           IF #statBatteryFamily1 = 16#0A THEN
               #HMI.State.Details.batFamily := 1;          //BAT1600
           ELSIF #statBatteryFamily1 = 16#09 THEN
               IF #statBatteryFamily2 = 16#07 THEN
                   #HMI.State.Details.batFamily := 3;          //Third Party Battery
               ELSE
                   #HMI.State.Details.batFamily := 2;          //UPS1100
               END_IF;
           END_IF;
           #HMI.State.batteryType := #statDataBatteryInfo.batteryDetails[0].batteryType;
           #HMI.State.endOfChargeVolt := INT_TO_REAL(#statDataBatteryInfo.batteryDetails[0].eocv) * 0.01;
           FOR #tempIterator := 0 TO 5 BY 1 DO
               #HMI.State.batteryDetails[#tempIterator].batteryLEDState := #statDataBatteryInfo.batteryDetails[#tempIterator].batLEDState;
               #HMI.State.batteryDetails[#tempIterator].batteryOpState := #statDataBatteryInfo.batteryDetails[#tempIterator].batOpState;
               #HMI.State.batteryDetails[#tempIterator].batteryCalcHealth := #statDataBatteryInfo.batteryDetails[#tempIterator].batCalcHealth;
           END_FOR;
           #HMI.State.chargingOpState := #statDataStateInfo.chargingOpState;
           // Cyclic Data
           #HMI.Mode.bufferMode := #statCyclicData[1];
           #HMI.Mode.readyForBuffering := #statCyclicData[2];
           #HMI.State.batteryChargeLevel := #statCyclicData[6];
           #statCyclicCount := 1;
       END_IF;

       //if Buffer_mode = 255, start Timer
       IF #HMI.Mode.bufferMode = 255 AND NOT #statBlockTimer AND NOT #statSetTimer THEN
           #statSetTimer := 1;
       END_IF;

       IF #HMI.Mode.bufferMode = 0 THEN
           #statSetTimer := 0;
           #statCmdDone := FALSE;
           #statBlockTimer := 0;
       END_IF;

       //BlockTimer - block
       #statTimerObj(IN := #statSetTimer,   // IN: BOOL
                     PT := #statBufferTime); // IN: TIME

       //Timer "Reset signal"
       IF #statTimerObj.Q = 1 THEN
           //if time elapse > UPS_ready_for_reset = 1
           #upsReadyForReset := 1;
           #statSetTimer := 0;
           #statBlockTimer := 1;
       END_IF;

       //reset UPS_ready_for_reset = 0 / set command parameter
       IF #upsExecuteReset = 1 AND NOT #statWrReq AND (#statBlockTimer = TRUE) AND (#statCmdDone = FALSE) THEN
           #statWrReq := 1;
           #statDataUPSCmd.commandID := 8207; //Command Remote Reset
           #statDataUPSCmd.parameter1 := INT_TO_BYTE(#statDataBufParam.bufferTime2);
           #statDataUPSCmd.parameter2 := #statDataResetParam;   //Parameter
           #upsReadyForReset := 0;
       END_IF;

       //write UPS Command
       #statDataRecordWrite(REQ := #statWrReq, ID := #addrIn, INDEX := 16, LEN := 4, RECORD := #statDataUPSCmd);

       IF #statDataRecordWrite.DONE OR #statDataRecordWrite.ERROR THEN
           #statWrReq := 0;
       END_IF;

       IF #statDataRecordWrite.DONE THEN
           #statCmdDone := TRUE;
       END_IF;

       // char to string > Order_number
       Chars_TO_Strg(Chars := #statDataDeviceInfo.orderNumber, pChars := 0, Cnt := 0, Strg => #statOrderNumberStr);
       #HMI.State.Details.orderNumber := #statOrderNumberStr;

       // char to string > Serial_number
       Chars_TO_Strg(Chars := #statDataDeviceInfo.serialNumber, pChars := 0, Cnt := 0, Strg => #statSerialNumberStr);
       #HMI.State.Details.serialNumber := #statSerialNumberStr;

       // char to string > Device_name
       Chars_TO_Strg(Chars := #statDataDeviceInfo.deviceName, pChars := 0, Cnt := 0, Strg => #statDeviceNameStr);
       #HMI.State.Details.deviceName := #statDeviceNameStr;

       // char to string > Version_number
       Chars_TO_Strg(Chars := #statDataDeviceInfo.versionNumber, pChars := 0, Cnt := 0, Strg => #statVersionNumberStr);
       #HMI.State.Details.versionNumber := #statVersionNumberStr;

       IF #statRetVal <> 0 AND #statCyclicCount = 1 THEN
           //setting acyclic data to default values
           #HMI.State.Details.orderNumber := ' ';
           #HMI.State.Details.serialNumber := ' ';
           #HMI.State.Details.deviceName := ' ';
           #HMI.State.Details.versionNumber := ' ';
           #HMI.State.Details.deviceHwRevision := 0;
           #HMI.State.Details.deviceSwRevision3 := 0;
           #HMI.State.Details.deviceSwRevision2 := 0;
           #HMI.State.Details.deviceSwRevision1 := 0;
           #HMI.State.numOfBatteries := 0;
           #HMI.State.Details.batFamily := 0;
           #HMI.State.batteryType := 0;
           #upsReadyForReset := 0;
       END_IF;
   END_IF;
END_REGION
END_FUNCTION_BLOCK

// folder: 1}Library/Analog

FUNCTION_BLOCK "Average"   // FB12, LAD
{ S7_Optimized_Access := 'TRUE' }
VERSION : 0.1
   VAR_INPUT
      TX1 : Real;
      TX2 : Real;
   END_VAR
   VAR_OUTPUT
      SAI : Real;
   END_VAR
BEGIN

REGION Network 1
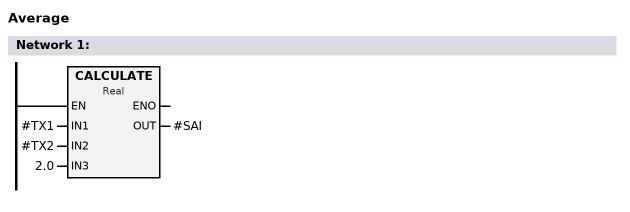
   RUNG wire#powerrail
      { S7_Templates := "SrcType := Real"; S7_Expression := "(IN1+IN2)/IN3" } Calculate(in1 := #TX1, in2 := #TX2, in3 := 2.0, out => #SAI)
   END_RUNG
   // the same network as SCL:
   #SAI := (#TX1+#TX2)/2.0;
END_REGION
END_FUNCTION_BLOCK

FUNCTION_BLOCK "AI Monitor"   // FB19, SCL
TITLE = Analog Input Monitor
{ S7_Optimized_Access := 'TRUE' }
AUTHOR : JLopez
VERSION : 0.1
// Monitor up to 6 Analog Inputs and execute AVG, in Range, deviation.
   VAR_INPUT
      "Enable Block" : Bool;   // Enable Block Execution
      "AI Num" : Int;   // Numbers of Analog Inputs Max: 6
      AvgSP : Real;   // Average SP Furnace Temperature
      "Min Range" : Real;   // Minimum Furnace Temperature Range
      "Max Range" : Real;   // Maximun Furnace Temperature Range
      MinAvgValue : Real := 0.0;   // Min Average Hysteresis Range
      MaxAvgValue : Real := 0.0;   // Max Average Hysteresis Range
      EnableDeviationMon : Bool;
      AlarmDeviation : Real := 25.0;
      MaxDeviation : Real := 50.0;   // Maximun deviation Allows
      MaxAboveTemp : Real := 50.0;
   END_VAR
   VAR_IN_OUT
      Avg : Real;   // Average Value
      AvgReached : Bool;   // Average Reached (Actual Average >=Avg-Minimum Average and <=Avg+Maximum Average
      AvgAlarm : Bool;
      ReadyToProcess : Bool;   // Conditions meet(Average,Range,Deviation) and ready to operate
      DeviationAlarm : Bool;
      DeviationFault : Bool;   // Deviation Fault Activated
      MaxAboveTempFault : Bool;   // Max Above Temperature Fault Activated
   END_VAR
   VAR
      AI_Mon : Struct
         InRange : Array[1..6] of Bool;   // TRUE=AI Ranges good, FALSE= AI Ranges not Good
         MinRange : Array[1..6] of Bool;   // TRUE=AI Minimun Range not Activated, False=AI Minimun Range Activated
         MaxRange : Array[1..6] of Bool;   // TRUE=AI Max Range not Activated, False=AI Max Range Activated
         Deviation : Array[1..6] of Bool;   // True= Analog Input Deviation; False=No Deviation
         DeviationAlarm : Array[1..6] of Bool;
         AboveTemp : Array[1..6] of Bool;   // Above Temperature Max Reached
      END_STRUCT;
      AI : Array[1..6] of Real;   // Analog Inputs
      AInputDeviation : Array[1..6] of Real;   // Actual Deviation Value between Analog Inputs
      AlarmsT : Struct
         DeviationAlarm : IEC_TIMER;
         DeviationFault : IEC_TIMER;
         MaxAbTempFault : IEC_TIMER;
      END_STRUCT;
      DeviationAlarmDelay : Time := T#5s;
      DeviationFaultDelay : Time := T#5s;
      MaxAboveTempFaultDelay : Time := T#5s;
      Aux : Struct
         DeviationAlarm : Bool;
         DeviationFault : Bool;
         MaxAboutTFault : Bool;
      END_STRUCT;
   END_VAR
   VAR_TEMP
      Indx : Int;
      TotalAIs : Real;   // Temporal Average
   END_VAR
BEGIN
   //**********Block description**********
   //The function of this block is to monitor the Analog inputs in the following way:
   //It has 3 presets; "AvgHysRanges"=Wish Average with a hysteresis value Min and Max, ex: Min=5, Max=5; will be consider that is in a good "Avg range" when is between this values. 
   //****************  "deviationValueSet"=Max Analog input(AI) Deviation between each other.
   //****************  "Min Range and Max Range"=Temperature Range of the Furnace that will be consider OK (Taking for each Analog Input).



   IF #"Enable Block" THEN

       IF #"AI Num" > 0 AND #"AI Num"<=6 AND #AvgSP>0.0  THEN  //"AI Num" is the quantity of Analog inputs to be monitor, should be less equal to 6 because 6 is the defined number as maximun (Block prepare to 6 Values).

           FOR #Indx := 1 TO #"AI Num" BY 1 DO     //Loop from index to "AI Num" parameter configured; Index will take values from 1,2,3..n when n="AI Num"
               #TotalAIs := #AI[#Indx] + #TotalAIs;  //Temporal Average Variable to be able to manipulate easly.

               #AI_Mon.MinRange[#Indx] := #AI[#Indx] > #"Min Range";   //Detect if each Analog Input is in Minimum Range, 1= AI in Range, 0= AI out of Range
               #AI_Mon.MaxRange[#Indx] := #AI[#Indx] < #"Max Range";   //Detect if each Analog Input is in Maximum Range, 1= AI in Range, 0= AI out of Range

                   IF #Indx>= #"AI Num"  THEN  //Condition to get the Avg to all the Analog Inputs.
                   #Avg := #TotalAIs / #"AI Num";  //Average of the total Analogs Inputs
                   END_IF;

                   #AI_Mon.InRange[#Indx] := #AI_Mon.MinRange[#Indx] AND #AI_Mon.MaxRange[#Indx]; //Analog Input in Range [Index].

                   IF #Indx < #"AI Num" THEN   //To avoid make the substraction of an AI that does not exist.
                       #AInputDeviation[#Indx] := #AI[#Indx] - #AI[#Indx + 1]; //Substract the AI[x]-AI[x+1]
                   ELSE    //To make the substraction from AI[6]-AI[1].
                       #AInputDeviation[#Indx] := #AI[#Indx] - #AI[#Indx - (#"AI Num"-1)];//Substract the AI[x]-AI[x+1]
                   END_IF;
                   #AInputDeviation[#Indx]:=ABS_REAL(#AInputDeviation[#Indx]); //Get the absolute value from the Substraction

                   IF #AInputDeviation[#Indx] > #AlarmDeviation THEN
                       #AI_Mon.DeviationAlarm[#Indx] := TRUE;  //There is a deviation Alarm between Temperatures (Analogs Inputs).
                   ELSE
                       #AI_Mon.DeviationAlarm[#Indx] := FALSE; //There is no deviation Alarm between Temperatures (Analogs Inputs)..
                   END_IF;

                   IF #AInputDeviation[#Indx] > #MaxDeviation THEN //If deviation is Higher that the preset
                       #AI_Mon.Deviation[#Indx] := TRUE;   //There a Max deviation between Temperatures (Analogs Inputs)..

                   ELSE
                       #AI_Mon.Deviation[#Indx] := FALSE;  //There is no deviation between Temperatures (Analogs Inputs)..

                   END_IF;
                   #AI_Mon.AboveTemp[#Indx] := #AI[#Indx] > (#AvgSP + #MaxAboveTemp);

               END_FOR;

               #AvgReached := #Avg >= (#AvgSP - #MinAvgValue) AND #Avg <= (#AvgSP + #MaxAvgValue);   //Hysteresis for the Average reached signal. 

               CASE #"AI Num" OF   //it will excecute depending of the quantity of Analogs Inputs that were configure in the "AI Num" Parameter.
               1:
                   IF #AI_Mon.InRange[1] AND #AvgReached THEN  //"1" Analog Input was set in the "AI Num" Parameter
                       #ReadyToProcess := TRUE;                //The Temperature is in the average.
                   ELSE
                       #ReadyToProcess := FALSE;               //The Temperature is not in the average.
                   END_IF;

               2:
                   IF #AI_Mon.InRange[1] AND #AI_Mon.InRange[2] AND #AvgReached THEN   //"2" Analog Inputs was set in the "AI Num" Parameter
                       #ReadyToProcess := TRUE;                //The Temperatures are in the average.
                   ELSE
                       #ReadyToProcess := FALSE;               //The Temperatures are not in the average.
                   END_IF;
               3:
                   IF #AI_Mon.InRange[1] AND #AI_Mon.InRange[2] AND #AI_Mon.InRange[3] AND #AvgReached THEN    //"3" Analog Inputs was set in the "AI Num" Parameter
                       #ReadyToProcess := TRUE;                //The Temperatures are in the average.
                   ELSE
                       #ReadyToProcess := FALSE;               //The Temperatures are not in the average.
                   END_IF;
               4:
                   IF #AI_Mon.InRange[1] AND #AI_Mon.InRange[2] AND #AI_Mon.InRange[3] AND #AI_Mon.InRange[4]
                       AND #AvgReached THEN     //"4" Analog Inputs was set in the "AI Num" Parameter
                       #ReadyToProcess := TRUE;                //The Temperatures are in the average.
                   ELSE
                       #ReadyToProcess := FALSE;               //The Temperatures are not in the average.
                   END_IF;
               5:
                   IF #AI_Mon.InRange[1] AND #AI_Mon.InRange[2] AND #AI_Mon.InRange[3] AND #AI_Mon.InRange[4]
                       AND #AI_Mon.InRange[5] AND #AvgReached THEN  //"5" Analog Inputs was set in the "AI Num" Parameter
                       #ReadyToProcess := TRUE;                //The Temperatures are in the average.
                   ELSE
                       #ReadyToProcess := FALSE;               //The Temperatures are not in the average.
                   END_IF;
               6:
                   IF #AI_Mon.InRange[1] AND #AI_Mon.InRange[2] AND #AI_Mon.InRange[3] AND #AI_Mon.InRange[4]
                       AND #AI_Mon.InRange[5] AND #AI_Mon.InRange[6] AND #AvgReached THEN   //"6" Analog Inputs was set in the "AI Num" Parameter
                       #ReadyToProcess := TRUE;                //The Temperatures are in the average.

                   ELSE
                       #ReadyToProcess := FALSE;               //The Temperatures are not in the average.
                   END_IF;
           END_CASE;

           IF #EnableDeviationMon THEN  //Deviation monitoring enable?
               //Deviation Alarm conditions
               IF #EnableDeviationMon AND (#AI_Mon.DeviationAlarm[1] OR #AI_Mon.DeviationAlarm[2]
                   OR #AI_Mon.DeviationAlarm[3] OR #AI_Mon.DeviationAlarm[4] OR #AI_Mon.DeviationAlarm[5] OR #AI_Mon.DeviationAlarm[6]) THEN
                   #Aux.DeviationAlarm := TRUE;
               ELSE
                   #Aux.DeviationAlarm := FALSE;
               END_IF;
               //Alarms Delay Timers
               #AlarmsT.DeviationAlarm.TON(IN := #Aux.DeviationAlarm,
                                           PT := #DeviationAlarmDelay);

               #DeviationAlarm := #AlarmsT.DeviationAlarm.Q;


               //Deviation Fault Conditions
               IF #EnableDeviationMon AND (#AI_Mon.Deviation[1] OR #AI_Mon.Deviation[2] OR #AI_Mon.Deviation[3]
                   OR #AI_Mon.Deviation[4] OR #AI_Mon.Deviation[5] OR #AI_Mon.Deviation[6]) THEN
                   #Aux.DeviationFault := TRUE;
               ELSE
                   #Aux.DeviationFault := FALSE;
               END_IF;
               //Alarms Delay Timers
               #AlarmsT.DeviationFault.TON(IN := #Aux.DeviationFault,
                                           PT := #DeviationFaultDelay);

               #DeviationFault := #AlarmsT.DeviationFault.Q;

               //Max Above Temp Fault Conditions
               IF #EnableDeviationMon AND (#AI_Mon.AboveTemp[1] OR #AI_Mon.AboveTemp[2] OR #AI_Mon.AboveTemp[3]
                   OR #AI_Mon.AboveTemp[4] OR #AI_Mon.AboveTemp[5] OR #AI_Mon.AboveTemp[6]) THEN
                   #Aux.MaxAboutTFault := TRUE;
               ELSE
                   #Aux.MaxAboutTFault := FALSE;
               END_IF;
               //Alarms Delay Timers
               #AlarmsT.MaxAbTempFault.TON(IN := #Aux.MaxAboutTFault,
                                           PT := #MaxAboveTempFaultDelay);

               #MaxAboveTempFault := #AlarmsT.MaxAbTempFault.Q;
           ELSE
               #DeviationAlarm := FALSE;
               #DeviationFault := FALSE;
               #MaxAboveTempFault := FALSE;
           END_IF;

       ELSE
           #Avg := 0.0;
           #ReadyToProcess := FALSE;
           #AvgReached := FALSE;
       END_IF;
   ELSE
       #Avg := 0.0;
       #ReadyToProcess := FALSE;
       #AvgReached := FALSE;
   END_IF;
END_FUNCTION_BLOCK

FUNCTION_BLOCK "AI Monitor_v2"   // FB20, SCL
TITLE = Analog Input Monitor
{ S7_Optimized_Access := 'TRUE' }
AUTHOR : JLopez
VERSION : 0.1
// Monitor up to 6 Analog Inputs and execute AVG, in Range, deviation.
   VAR_INPUT
      "Enable Block" : Bool;   // Enable Block Execution
      "AI Num" : Int;   // Numbers of Analog Inputs Max: 6
      AvgSP : Real;   // Average SP Furnace Temperature
      "Min Range" : Real;   // Minimum Furnace Temperature Range
      "Max Range" : Real;   // Maximun Furnace Temperature Range
      MinAvgValue : Real := 0.0;   // Min Average Hysteresis Range
      MaxAvgValue : Real := 0.0;   // Max Average Hysteresis Range
      EnableDeviationMon : Bool;
      AlarmDeviation : Real := 25.0;
      MaxDeviation : Real := 50.0;   // Maximun deviation Allows
      MaxAboveTemp : Real := 50.0;
   END_VAR
   VAR_IN_OUT
      Avg : Real;   // Average Value
      AvgReached : Bool;   // Average Reached (Actual Average >=Avg-Minimum Average and <=Avg+Maximum Average
      AvgAlarm : Bool;
      ReadyToProcess : Bool;   // Conditions meet(Average,Range,Deviation) and ready to operate
      DeviationAlarm : Bool;
      DeviationFault : Bool;   // Deviation Fault Activated
      MaxAboveTempFault : Bool;   // Max Above Temperature Fault Activated
   END_VAR
   VAR
      AI_Mon : Struct
         InRange : Array[1..6] of Bool;   // TRUE=AI Ranges good, FALSE= AI Ranges not Good
         MinRange : Array[1..6] of Bool;   // TRUE=AI Minimun Range not Activated, False=AI Minimun Range Activated
         MaxRange : Array[1..6] of Bool;   // TRUE=AI Max Range not Activated, False=AI Max Range Activated
         Deviation : Array[1..6, 1..6] of Bool;   // True= Analog Input Deviation; False=No Deviation
         DeviationAlarm : Array[1..6, 1..6] of Bool;
         AboveTemp : Array[1..6] of Bool;   // Above Temperature Max Reached
      END_STRUCT;
      AI : Array[1..6] of Real;   // Analog Inputs
      AInputDeviation : Array[1..6, 1..6] of Real;   // Actual Deviation Value between Analog Inputs
      AlarmsT : Struct
         DeviationAlarm : IEC_TIMER;
         DeviationFault : IEC_TIMER;
         MaxAbTempFault : IEC_TIMER;
      END_STRUCT;
      DeviationAlarmDelay : Time := T#5s;
      DeviationFaultDelay : Time := T#5s;
      MaxAboveTempFaultDelay : Time := T#5s;
      Aux : Struct
         DeviationAlarm : Bool;
         DeviationFault : Bool;
         MaxAboutTFault : Bool;
      END_STRUCT;
   END_VAR
   VAR_TEMP
      DeviationAlarmActivated : Bool;
      DeviationFaultActivated : Bool;
      Indx : Int;
      Indx2 : Int;
      TotalAIs : Real;   // Temporal Average
   END_VAR
BEGIN
   //**********Block description**********
   //The function of this block is to monitor the Analog inputs in the following way:
   //It has 3 presets; "AvgHysRanges"=Wish Average with a hysteresis value Min and Max, ex: Min=5, Max=5; will be consider that is in a good "Avg range" when is between this values. 
   //****************  "deviationValueSet"=Max Analog input(AI) Deviation between each other.
   //****************  "Min Range and Max Range"=Temperature Range of the Furnace that will be consider OK (Taking for each Analog Input).



   IF #"Enable Block" THEN

       IF #"AI Num" > 0 AND #"AI Num"<=6 AND #AvgSP>0.0  THEN  //"AI Num" is the quantity of Analog inputs to be monitor, should be less equal to 6 because 6 is the defined number as maximun (Block prepare to 6 Values).

           FOR #Indx := 1 TO #"AI Num" BY 1 DO     //Loop from index to "AI Num" parameter configured; Index will take values from 1,2,3..n when n="AI Num"
               #TotalAIs := #AI[#Indx] + #TotalAIs;  //Temporal Average Variable to be able to manipulate easly.

               #AI_Mon.MinRange[#Indx] := #AI[#Indx] > #"Min Range";   //Detect if each Analog Input is in Minimum Range, 1= AI in Range, 0= AI out of Range
               #AI_Mon.MaxRange[#Indx] := #AI[#Indx] < #"Max Range";   //Detect if each Analog Input is in Maximum Range, 1= AI in Range, 0= AI out of Range

                   IF #Indx>= #"AI Num"  THEN  //Condition to get the Avg to all the Analog Inputs.
                   #Avg := #TotalAIs / #"AI Num";  //Average of the total Analogs Inputs
                   END_IF;

                   #AI_Mon.InRange[#Indx] := #AI_Mon.MinRange[#Indx] AND #AI_Mon.MaxRange[#Indx]; //Analog Input in Range [Index].

                   //Loop for calculate the deviation of the AIs
                   FOR #Indx2 := 1 TO #"AI Num" BY 1 DO

                       IF #Indx2 < #"AI Num" THEN   //To avoid make the substraction of an AI that does not exist.
                           #AInputDeviation[#Indx, #Indx2] := #AI[#Indx2] - #AI[#Indx2 + 1]; //Substract the AI[x]-AI[x+1]
                       ELSE    //To make the substraction from AI[6]-AI[1].
                           #AInputDeviation[#Indx, #Indx2] := #AI[#Indx2] - #AI[#Indx2 - (#"AI Num" - 1)];//Substract the AI[x]-AI[x+1]
                       END_IF;

                       #AInputDeviation[#Indx,#Indx2] := ABS_REAL(#AInputDeviation[#Indx,#Indx2]); //Get the absolute value from the Substraction

                       IF #AInputDeviation[#Indx,#Indx2] > #AlarmDeviation THEN
                           #AI_Mon.DeviationAlarm[#Indx,#Indx2] := TRUE;  //There is a deviation Alarm between Temperatures (Analogs Inputs).
                           #DeviationAlarmActivated := TRUE;
                       ELSE
                           #AI_Mon.DeviationAlarm[#Indx,#Indx2] := FALSE; //There is no deviation Alarm between Temperatures (Analogs Inputs)..

                       END_IF;

                       IF #AInputDeviation[#Indx,#Indx2] > #MaxDeviation THEN //If deviation is Higher that the preset
                           #AI_Mon.Deviation[#Indx,#Indx2] := TRUE;   //There a Max deviation between Temperatures (Analogs Inputs)..
                           #DeviationFaultActivated := TRUE;
                       ELSE
                           #AI_Mon.Deviation[#Indx,#Indx2] := FALSE;  //There is no deviation between Temperatures (Analogs Inputs)..

                       END_IF;
                   END_FOR;

                   #AI_Mon.AboveTemp[#Indx] := #AI[#Indx] > (#AvgSP + #MaxAboveTemp);

               END_FOR;

               #AvgReached := #Avg >= (#AvgSP - #MinAvgValue) AND #Avg <= (#AvgSP + #MaxAvgValue);   //Hysteresis for the Average reached signal. 

               CASE #"AI Num" OF   //it will excecute depending of the quantity of Analogs Inputs that were configure in the "AI Num" Parameter.
               1:
                   IF #AI_Mon.InRange[1] AND #AvgReached THEN  //"1" Analog Input was set in the "AI Num" Parameter
                       #ReadyToProcess := TRUE;                //The Temperature is in the average.
                   ELSE
                       #ReadyToProcess := FALSE;               //The Temperature is not in the average.
                   END_IF;

               2:
                   IF #AI_Mon.InRange[1] AND #AI_Mon.InRange[2] AND #AvgReached THEN   //"2" Analog Inputs was set in the "AI Num" Parameter
                       #ReadyToProcess := TRUE;                //The Temperatures are in the average.
                   ELSE
                       #ReadyToProcess := FALSE;               //The Temperatures are not in the average.
                   END_IF;
               3:
                   IF #AI_Mon.InRange[1] AND #AI_Mon.InRange[2] AND #AI_Mon.InRange[3] AND #AvgReached THEN    //"3" Analog Inputs was set in the "AI Num" Parameter
                       #ReadyToProcess := TRUE;                //The Temperatures are in the average.
                   ELSE
                       #ReadyToProcess := FALSE;               //The Temperatures are not in the average.
                   END_IF;
               4:
                   IF #AI_Mon.InRange[1] AND #AI_Mon.InRange[2] AND #AI_Mon.InRange[3] AND #AI_Mon.InRange[4]
                       AND #AvgReached THEN     //"4" Analog Inputs was set in the "AI Num" Parameter
                       #ReadyToProcess := TRUE;                //The Temperatures are in the average.
                   ELSE
                       #ReadyToProcess := FALSE;               //The Temperatures are not in the average.
                   END_IF;
               5:
                   IF #AI_Mon.InRange[1] AND #AI_Mon.InRange[2] AND #AI_Mon.InRange[3] AND #AI_Mon.InRange[4]
                       AND #AI_Mon.InRange[5] AND #AvgReached THEN  //"5" Analog Inputs was set in the "AI Num" Parameter
                       #ReadyToProcess := TRUE;                //The Temperatures are in the average.
                   ELSE
                       #ReadyToProcess := FALSE;               //The Temperatures are not in the average.
                   END_IF;
               6:
                   IF #AI_Mon.InRange[1] AND #AI_Mon.InRange[2] AND #AI_Mon.InRange[3] AND #AI_Mon.InRange[4]
                       AND #AI_Mon.InRange[5] AND #AI_Mon.InRange[6] AND #AvgReached THEN   //"6" Analog Inputs was set in the "AI Num" Parameter
                       #ReadyToProcess := TRUE;                //The Temperatures are in the average.

                   ELSE
                       #ReadyToProcess := FALSE;               //The Temperatures are not in the average.
                   END_IF;
           END_CASE;

           IF #EnableDeviationMon THEN  //Deviation monitoring enable?
               //Deviation Alarm conditions
               IF #EnableDeviationMon AND #DeviationAlarmActivated THEN
                   #Aux.DeviationAlarm := TRUE;
               ELSE
                   #Aux.DeviationAlarm := FALSE;
               END_IF;
               //Alarms Delay Timers
               #AlarmsT.DeviationAlarm.TON(IN := #Aux.DeviationAlarm,
                                           PT := #DeviationAlarmDelay);

               #DeviationAlarm := #AlarmsT.DeviationAlarm.Q;


               //Deviation Fault Conditions
               IF #EnableDeviationMon AND #DeviationFaultActivated THEN
                   #Aux.DeviationFault := TRUE;
               ELSE
                   #Aux.DeviationFault := FALSE;
               END_IF;
               //Alarms Delay Timers
               #AlarmsT.DeviationFault.TON(IN := #Aux.DeviationFault,
                                           PT := #DeviationFaultDelay);

               #DeviationFault := #AlarmsT.DeviationFault.Q;

               //Max Above Temp Fault Conditions
               IF #EnableDeviationMon AND (#AI_Mon.AboveTemp[1] OR #AI_Mon.AboveTemp[2] OR #AI_Mon.AboveTemp[3]
                   OR #AI_Mon.AboveTemp[4] OR #AI_Mon.AboveTemp[5] OR #AI_Mon.AboveTemp[6]) THEN
                   #Aux.MaxAboutTFault := TRUE;
               ELSE
                   #Aux.MaxAboutTFault := FALSE;
               END_IF;
               //Alarms Delay Timers
               #AlarmsT.MaxAbTempFault.TON(IN := #Aux.MaxAboutTFault,
                                           PT := #MaxAboveTempFaultDelay);

               #MaxAboveTempFault := #AlarmsT.MaxAbTempFault.Q;
           ELSE
               #DeviationAlarm := FALSE;
               #DeviationFault := FALSE;
               #MaxAboveTempFault := FALSE;
           END_IF;

       ELSE
           #Avg := 0.0;
           #ReadyToProcess := FALSE;
           #AvgReached := FALSE;
       END_IF;
   ELSE
       #Avg := 0.0;
       #ReadyToProcess := FALSE;
       #AvgReached := FALSE;
   END_IF;
END_FUNCTION_BLOCK

FUNCTION_BLOCK "3 Analog Voting"   // FB66, LAD
{ S7_Optimized_Access := 'TRUE' }
VERSION : 0.1
   VAR_INPUT
      analog1 : Real;   // Scaled Value 1
      analog2 : Real;   // Scale Value 2
      analog3 : Real;   // Scaled Value 3
      fault1 : Bool;   // Fault of Transmitter 1
      fault2 : Bool;   // Fault of Transmitter 2
      fault3 : Bool;   // Fault of Transmitter 3
   END_VAR
   VAR_OUTPUT
      activeValue : Real;   // value selected to be Output (median, lowest, highest, average, only one)
      medianValue : Real;   // Value Selected by operator
      masterTrip : Bool;   // 2oo3 voting (deviation, lowlow, highhigh, wirebreak) mixed
      masterTripLowLow : Bool;   // 2oo3 voting (deviation, lowlow,wirebreak) mixed
      masterTripHighHigh : Bool;   // 2oo3 voting (deviation, highhigh, wirebreak) mixed
      HHT : Bool;   // HH trip voting
      HT : Bool;   // H trip voting
      LT : Bool;   // L trip voting
      LLT : Bool;   // LL trip voting
   END_VAR
   VAR
      HMI : Struct
         Config : Struct
            deviationTolerance : Real := 30.0;
            Limits : Struct
               HH : Real := 100.0;
               H : Real := 80.0;
               L : Real := 20.0;
               LL : Real := 10.0;
            END_STRUCT;
         END_STRUCT;
         Control : Struct
            mode : Int := 5;
            failMode : Int := 4;
         END_STRUCT;
         Alarms : Struct
            "HH Value 1" : Bool;
            "HH Value 2" : Bool;
            "HH Value 3" : Bool;
            "H Value 1" : Bool;
            "H Value 2" : Bool;
            "H Value 3" : Bool;
            "L Value 1" : Bool;
            "L Value 2" : Bool;
            "L Value 3" : Bool;
            "LL Value 1" : Bool;
            "LL Value 2" : Bool;
            "LL Value 3" : Bool;
            "Value 1 Deviation" : Bool;
            "Value 2 Deviation" : Bool;
            "Value 3 Deviation" : Bool;
            deviationGeneralAlarm : Bool;
            activeValueHH : Bool;
            activeValueH : Bool;
            activeValueL : Bool;
            acrtiveValueLL : Bool;
            oneTxFaulted : Bool;
            twoTxFaulted : Bool;
            triggers : Array[0..15] of Bool;
         END_STRUCT;
      END_STRUCT;
      "HH Vote 1" : "HLR";
      "HH Vote 2" : "HLR";
      "HH Vote 3" : "HLR";
      "HH Vote activeValue" : "HLR";
      "H Vote 1" : "HLR";
      "H Vote 2" : "HLR";
      "H Vote 3" : "HLR";
      "H Vote activeValue" : "HLR";
      "L Vote 1" : "LLR";
      "L Vote 2" : "LLR";
      "L Vote 3" : "LLR";
      "L Vote activeValue" : "LLR";
      "LL Vote 1" : "LLR";
      "LL Vote 2" : "LLR";
      "LL Vote 3" : "LLR";
      "LL Vote activeValue" : "LLR";
      value1Deviated : Bool;
      value2Deviated : Bool;
      value3Deviated : Bool;
   END_VAR
   VAR_TEMP
      N1 : Real;
      AN1 : Real;
      N2 : Real;
      AN2 : Real;
      N3 : Real;
      AN3 : Real;
      average : Real;
      highest : Real;
      lowest : Real;
      tempMedian : Real;
   END_VAR
   VAR_TEMP   // added for the SCL form of the ladder/FBD networks
      _w1 : Bool;
   END_VAR
BEGIN

REGION Network 1: Transmitter failure
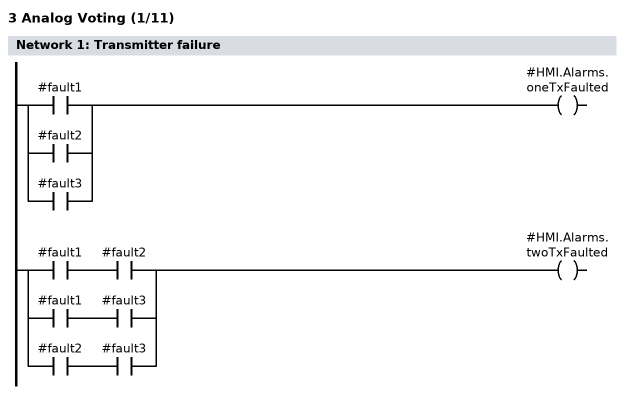
   RUNG wire#powerrail
      Contact( #fault1 )
      wire#w1
      Coil( #HMI.Alarms.oneTxFaulted )
   END_RUNG
   RUNG wire#powerrail
      Contact( #fault2 )
   END_RUNG wire#w1
   RUNG wire#powerrail
      Contact( #fault3 )
   END_RUNG wire#w1
   RUNG wire#powerrail
      Contact( #fault1 )
      Contact( #fault2 )
      wire#w2
      Coil( #HMI.Alarms.twoTxFaulted )
   END_RUNG
   RUNG wire#powerrail
      Contact( #fault1 )
      Contact( #fault3 )
   END_RUNG wire#w2
   RUNG wire#powerrail
      Contact( #fault2 )
      Contact( #fault3 )
   END_RUNG wire#w2
   // the same network as SCL:
   #HMI.Alarms.oneTxFaulted := #fault1 OR #fault2 OR #fault3;
   #HMI.Alarms.twoTxFaulted := (#fault1 AND #fault2) OR (#fault1 AND #fault3) OR (#fault2 AND #fault3);
END_REGION

REGION Network 2: HighestLowest
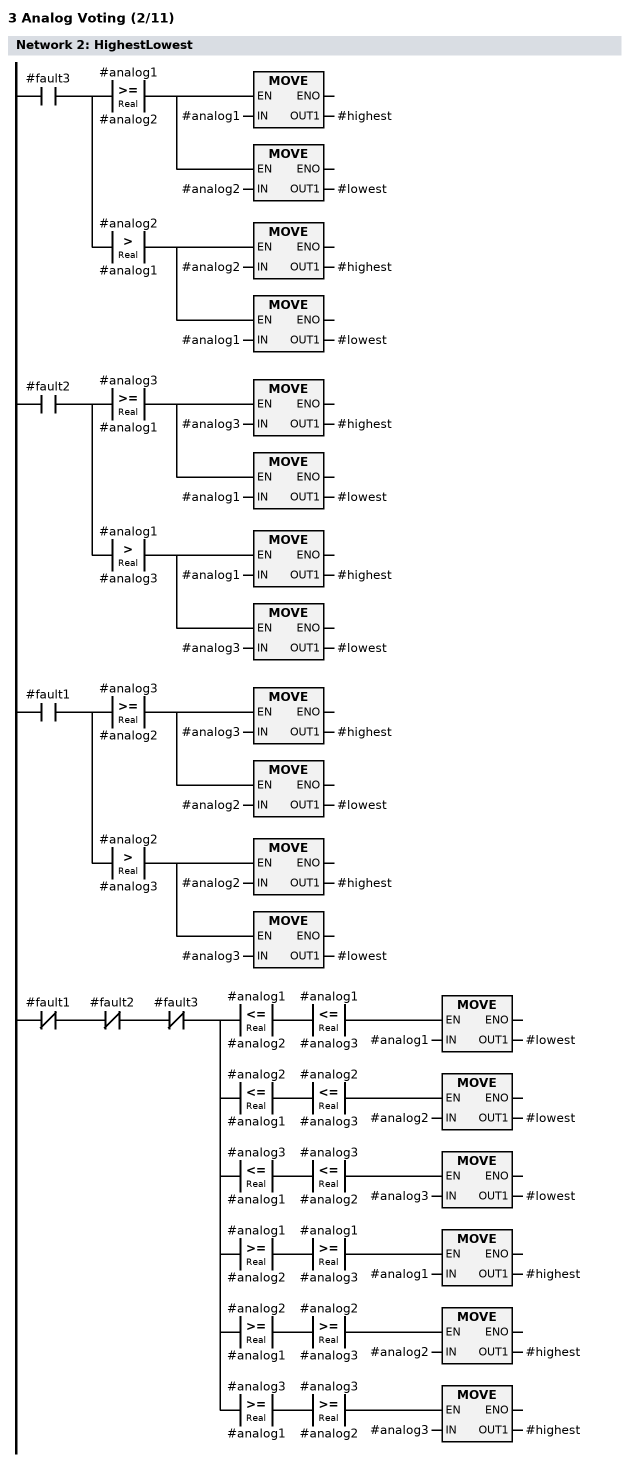
   RUNG wire#powerrail
      Contact( #fault3 )
      wire#w1
      { S7_Templates := "SrcType := Real" } GE_Contact(in1 := #analog1, in2 := #analog2)
      wire#w2
      Move(in := #analog1, out1 => #highest)
   END_RUNG
   RUNG wire#w2
      Move(in := #analog2, out1 => #lowest)
   END_RUNG
   RUNG wire#w1
      { S7_Templates := "SrcType := Real" } GT_Contact(in1 := #analog2, in2 := #analog1)
      wire#w3
      Move(in := #analog2, out1 => #highest)
   END_RUNG
   RUNG wire#w3
      Move(in := #analog1, out1 => #lowest)
   END_RUNG
   RUNG wire#powerrail
      Contact( #fault2 )
      wire#w4
      { S7_Templates := "SrcType := Real" } GE_Contact(in1 := #analog3, in2 := #analog1)
      wire#w5
      Move(in := #analog3, out1 => #highest)
   END_RUNG
   RUNG wire#w5
      Move(in := #analog1, out1 => #lowest)
   END_RUNG
   RUNG wire#w4
      { S7_Templates := "SrcType := Real" } GT_Contact(in1 := #analog1, in2 := #analog3)
      wire#w6
      Move(in := #analog1, out1 => #highest)
   END_RUNG
   RUNG wire#w6
      Move(in := #analog3, out1 => #lowest)
   END_RUNG
   RUNG wire#powerrail
      Contact( #fault1 )
      wire#w7
      { S7_Templates := "SrcType := Real" } GE_Contact(in1 := #analog3, in2 := #analog2)
      wire#w8
      Move(in := #analog3, out1 => #highest)
   END_RUNG
   RUNG wire#w8
      Move(in := #analog2, out1 => #lowest)
   END_RUNG
   RUNG wire#w7
      { S7_Templates := "SrcType := Real" } GT_Contact(in1 := #analog2, in2 := #analog3)
      wire#w9
      Move(in := #analog2, out1 => #highest)
   END_RUNG
   RUNG wire#w9
      Move(in := #analog3, out1 => #lowest)
   END_RUNG
   RUNG wire#powerrail
      I_Contact( #fault1 )
      I_Contact( #fault2 )
      I_Contact( #fault3 )
      wire#w10
      { S7_Templates := "SrcType := Real" } LE_Contact(in1 := #analog1, in2 := #analog2)
      { S7_Templates := "SrcType := Real" } LE_Contact(in1 := #analog1, in2 := #analog3)
      Move(in := #analog1, out1 => #lowest)
   END_RUNG
   RUNG wire#w10
      { S7_Templates := "SrcType := Real" } LE_Contact(in1 := #analog2, in2 := #analog1)
      { S7_Templates := "SrcType := Real" } LE_Contact(in1 := #analog2, in2 := #analog3)
      Move(in := #analog2, out1 => #lowest)
   END_RUNG
   RUNG wire#w10
      { S7_Templates := "SrcType := Real" } LE_Contact(in1 := #analog3, in2 := #analog1)
      { S7_Templates := "SrcType := Real" } LE_Contact(in1 := #analog3, in2 := #analog2)
      Move(in := #analog3, out1 => #lowest)
   END_RUNG
   RUNG wire#w10
      { S7_Templates := "SrcType := Real" } GE_Contact(in1 := #analog1, in2 := #analog2)
      { S7_Templates := "SrcType := Real" } GE_Contact(in1 := #analog1, in2 := #analog3)
      Move(in := #analog1, out1 => #highest)
   END_RUNG
   RUNG wire#w10
      { S7_Templates := "SrcType := Real" } GE_Contact(in1 := #analog2, in2 := #analog1)
      { S7_Templates := "SrcType := Real" } GE_Contact(in1 := #analog2, in2 := #analog3)
      Move(in := #analog2, out1 => #highest)
   END_RUNG
   RUNG wire#w10
      { S7_Templates := "SrcType := Real" } GE_Contact(in1 := #analog3, in2 := #analog1)
      { S7_Templates := "SrcType := Real" } GE_Contact(in1 := #analog3, in2 := #analog2)
      Move(in := #analog3, out1 => #highest)
   END_RUNG
   // the same network as SCL:
   IF #fault3 AND (#analog1 >= #analog2) THEN
       #highest := #analog1;
       #lowest := #analog2;
   END_IF;
   IF #fault3 AND (#analog2 > #analog1) THEN
       #highest := #analog2;
       #lowest := #analog1;
   END_IF;
   IF #fault2 AND (#analog3 >= #analog1) THEN
       #highest := #analog3;
       #lowest := #analog1;
   END_IF;
   IF #fault2 AND (#analog1 > #analog3) THEN
       #highest := #analog1;
       #lowest := #analog3;
   END_IF;
   IF #fault1 AND (#analog3 >= #analog2) THEN
       #highest := #analog3;
       #lowest := #analog2;
   END_IF;
   IF #fault1 AND (#analog2 > #analog3) THEN
       #highest := #analog2;
       #lowest := #analog3;
   END_IF;
   #_w1 := NOT #fault1 AND NOT #fault2 AND NOT #fault3;
   IF #_w1 AND (#analog1 <= #analog2) AND (#analog1 <= #analog3) THEN #lowest := #analog1; END_IF;
   IF #_w1 AND (#analog2 <= #analog1) AND (#analog2 <= #analog3) THEN #lowest := #analog2; END_IF;
   IF #_w1 AND (#analog3 <= #analog1) AND (#analog3 <= #analog2) THEN #lowest := #analog3; END_IF;
   IF #_w1 AND (#analog1 >= #analog2) AND (#analog1 >= #analog3) THEN #highest := #analog1; END_IF;
   IF #_w1 AND (#analog2 >= #analog1) AND (#analog2 >= #analog3) THEN #highest := #analog2; END_IF;
   IF #_w1 AND (#analog3 >= #analog1) AND (#analog3 >= #analog2) THEN #highest := #analog3; END_IF;
END_REGION

REGION Network 3: Two Transmitters Failed...select last value
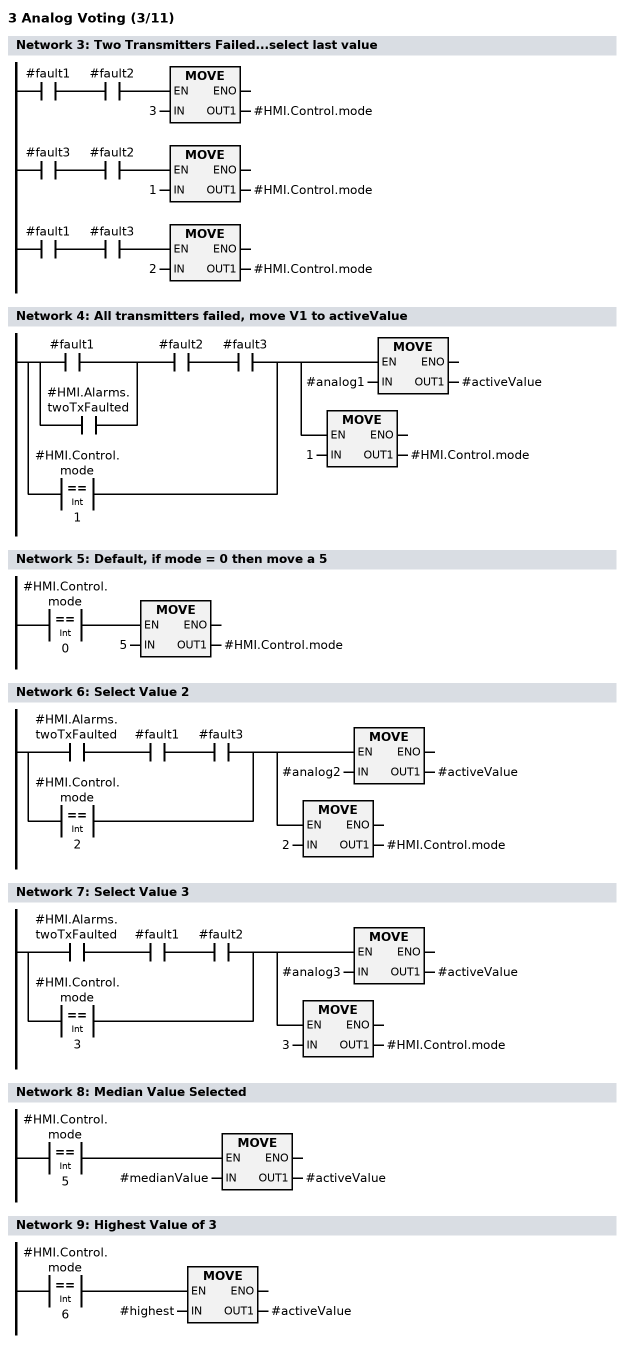
   RUNG wire#powerrail
      Contact( #fault1 )
      Contact( #fault2 )
      Move(in := 3, out1 => #HMI.Control.mode)
   END_RUNG
   RUNG wire#powerrail
      Contact( #fault3 )
      Contact( #fault2 )
      Move(in := 1, out1 => #HMI.Control.mode)
   END_RUNG
   RUNG wire#powerrail
      Contact( #fault1 )
      Contact( #fault3 )
      Move(in := 2, out1 => #HMI.Control.mode)
   END_RUNG
   // the same network as SCL:
   IF #fault1 AND #fault2 THEN #HMI.Control.mode := 3; END_IF;
   IF #fault3 AND #fault2 THEN #HMI.Control.mode := 1; END_IF;
   IF #fault1 AND #fault3 THEN #HMI.Control.mode := 2; END_IF;
END_REGION

REGION Network 4: All transmitters failed, move V1 to activeValue
   RUNG wire#powerrail
      Contact( #fault1 )
      wire#w1
      Contact( #fault2 )
      Contact( #fault3 )
      wire#w2
      Move(in := #analog1, out1 => #activeValue)
   END_RUNG
   RUNG wire#powerrail
      Contact( #HMI.Alarms.twoTxFaulted )
   END_RUNG wire#w1
   RUNG wire#powerrail
      { S7_Templates := "SrcType := Int" } EQ_Contact(in1 := #HMI.Control.mode, in2 := 1)
   END_RUNG wire#w2
   RUNG wire#w2
      Move(in := 1, out1 => #HMI.Control.mode)
   END_RUNG
   // the same network as SCL:
   IF ((#fault1 OR #HMI.Alarms.twoTxFaulted) AND #fault2 AND #fault3) OR (#HMI.Control.mode = 1) THEN
       #activeValue := #analog1;
       #HMI.Control.mode := 1;
   END_IF;
END_REGION

REGION Network 5: Default, if mode = 0 then move a 5
   RUNG wire#powerrail
      { S7_Templates := "SrcType := Int" } EQ_Contact(in1 := #HMI.Control.mode, in2 := 0)
      Move(in := 5, out1 => #HMI.Control.mode)
   END_RUNG
   // the same network as SCL:
   IF #HMI.Control.mode = 0 THEN #HMI.Control.mode := 5; END_IF;
END_REGION

REGION Network 6: Select Value 2
   RUNG wire#powerrail
      Contact( #HMI.Alarms.twoTxFaulted )
      Contact( #fault1 )
      Contact( #fault3 )
      wire#w1
      Move(in := #analog2, out1 => #activeValue)
   END_RUNG
   RUNG wire#powerrail
      { S7_Templates := "SrcType := Int" } EQ_Contact(in1 := #HMI.Control.mode, in2 := 2)
   END_RUNG wire#w1
   RUNG wire#w1
      Move(in := 2, out1 => #HMI.Control.mode)
   END_RUNG
   // the same network as SCL:
   IF (#HMI.Alarms.twoTxFaulted AND #fault1 AND #fault3) OR (#HMI.Control.mode = 2) THEN
       #activeValue := #analog2;
       #HMI.Control.mode := 2;
   END_IF;
END_REGION

REGION Network 7: Select Value 3
   RUNG wire#powerrail
      Contact( #HMI.Alarms.twoTxFaulted )
      Contact( #fault1 )
      Contact( #fault2 )
      wire#w1
      Move(in := #analog3, out1 => #activeValue)
   END_RUNG
   RUNG wire#powerrail
      { S7_Templates := "SrcType := Int" } EQ_Contact(in1 := #HMI.Control.mode, in2 := 3)
   END_RUNG wire#w1
   RUNG wire#w1
      Move(in := 3, out1 => #HMI.Control.mode)
   END_RUNG
   // the same network as SCL:
   IF (#HMI.Alarms.twoTxFaulted AND #fault1 AND #fault2) OR (#HMI.Control.mode = 3) THEN
       #activeValue := #analog3;
       #HMI.Control.mode := 3;
   END_IF;
END_REGION

REGION Network 8: Median Value Selected
   RUNG wire#powerrail
      { S7_Templates := "SrcType := Int" } EQ_Contact(in1 := #HMI.Control.mode, in2 := 5)
      Move(in := #medianValue, out1 => #activeValue)
   END_RUNG
   // the same network as SCL:
   IF #HMI.Control.mode = 5 THEN #activeValue := #medianValue; END_IF;
END_REGION

REGION Network 9: Highest Value of 3
   RUNG wire#powerrail
      { S7_Templates := "SrcType := Int" } EQ_Contact(in1 := #HMI.Control.mode, in2 := 6)
      Move(in := #highest, out1 => #activeValue)
   END_RUNG
   // the same network as SCL:
   IF #HMI.Control.mode = 6 THEN #activeValue := #highest; END_IF;
END_REGION

REGION Network 10: Lowest Value of 3
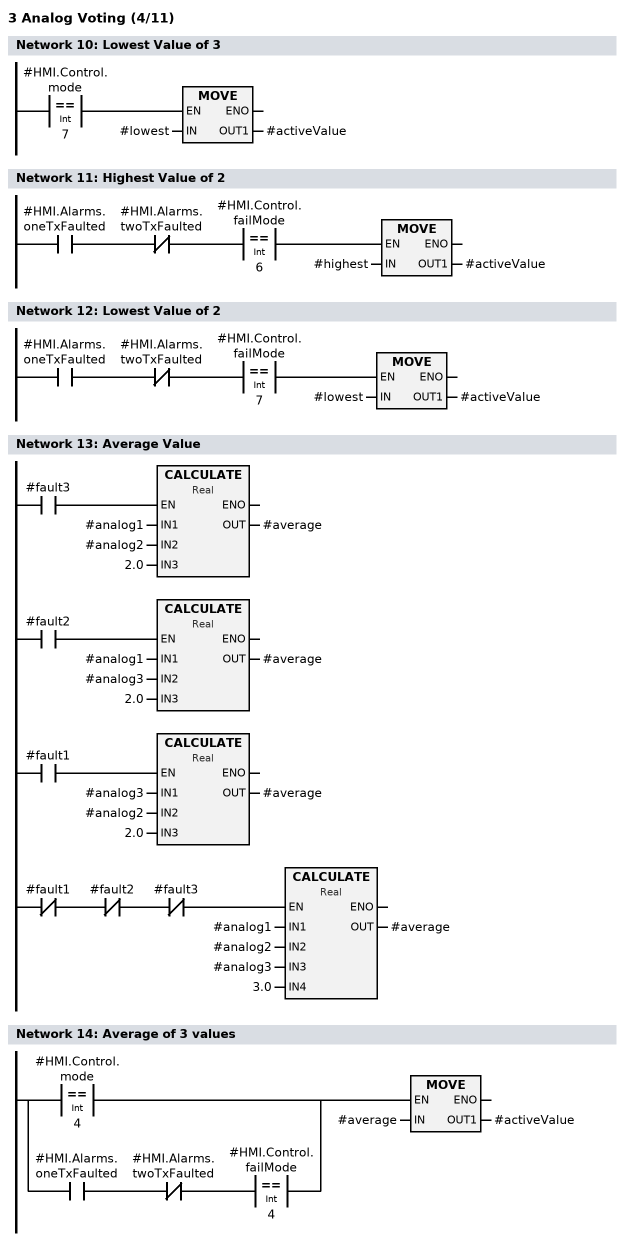
   RUNG wire#powerrail
      { S7_Templates := "SrcType := Int" } EQ_Contact(in1 := #HMI.Control.mode, in2 := 7)
      Move(in := #lowest, out1 => #activeValue)
   END_RUNG
   // the same network as SCL:
   IF #HMI.Control.mode = 7 THEN #activeValue := #lowest; END_IF;
END_REGION

REGION Network 11: Highest Value of 2
   RUNG wire#powerrail
      Contact( #HMI.Alarms.oneTxFaulted )
      I_Contact( #HMI.Alarms.twoTxFaulted )
      { S7_Templates := "SrcType := Int" } EQ_Contact(in1 := #HMI.Control.failMode, in2 := 6)
      Move(in := #highest, out1 => #activeValue)
   END_RUNG
   // the same network as SCL:
   IF #HMI.Alarms.oneTxFaulted AND NOT #HMI.Alarms.twoTxFaulted AND (#HMI.Control.failMode = 6) THEN
       #activeValue := #highest;
   END_IF;
END_REGION
